(* Logix 5000 project; controller FV vendor 1 type 14 code 217 rev 31.11; software revision 31.00; part 50 of 63 *)
(* tags used below, declared in another part *)
   CheckTimeMask : INT;
   Delphi_Does_Eng_Func : BOOL;
   FV_ALARM : PlantItem;   // ALARM
   FV_AV1 : PlantItem;   // AV1
   FV_AV1A : PlantItem;   // AV1A
   FV_AV2 : PlantItem;   // AV2
   FV_AV3 : PlantItem;   // AV3
   FV_AV4 : PlantItem;   // AV4
   FV_AV4A : PlantItem;   // AV4A
   FV_FV10C : PlantItem;   // FV10C
   FV_FV10J : PlantItem;   // FV10J
   FV_FV11C : PlantItem;   // FV11C
   FV_FV11J : PlantItem;   // FV11J
   FV_FV12C : PlantItem;   // FV12C
   FV_FV12J : PlantItem;   // FV12J
   FV_FV13C : PlantItem;   // FV13C
   FV_FV13J : PlantItem;   // FV13J
   FV_FV14C : PlantItem;   // FV14C
   FV_FV14J : PlantItem;   // FV14J
   FV_FV15C : PlantItem;   // FV15C
   FV_FV15J : PlantItem;   // FV15J
   FV_FV16C : PlantItem;   // FV16C
   FV_FV16J : PlantItem;   // FV16J
   FV_FV17C : PlantItem;   // FV17C
   FV_FV17J : PlantItem;   // FV17J
   FV_FV18C : PlantItem;   // FV18C
   FV_FV18J : PlantItem;   // FV18J
   FV_FV19C : PlantItem;   // FV19C
   FV_FV19J : PlantItem;   // FV19J
   FV_FV20C : PlantItem;   // FV20C
   FV_FV20J : PlantItem;   // FV20J
   FV_FV21C : PlantItem;   // FV21C
   FV_FV21J : PlantItem;   // FV21J
   FV_FV22C : PlantItem;   // FV22C
   FV_FV22J : PlantItem;   // FV22J
   FV_FV23C : PlantItem;   // FV23C
   FV_FV23J : PlantItem;   // FV23J
   FV_FV24C : PlantItem;   // FV24C
   FV_FV24J : PlantItem;   // FV24J
   FV_FV25C : PlantItem;   // FV25C
   FV_FV25J : PlantItem;   // FV25J
   FV_FV26C : PlantItem;   // FV26C
   FV_FV26J : PlantItem;   // FV26J
   FV_FV27C : PlantItem;   // FV27C
   FV_FV27J : PlantItem;   // FV27J
   FV_FV28C : PlantItem;   // FV28C
   FV_FV28J : PlantItem;   // FV28J
   FV_FV29C : PlantItem;   // FV29C
   FV_FV29J : PlantItem;   // FV29J
   FV_FV30C : PlantItem;   // FV30C
   FV_FV30J : PlantItem;   // FV30J
   FV_FV31C : PlantItem;   // FV31C
   FV_FV31J : PlantItem;   // FV31J
   FV_N255 : INT[255];   // Old Checkwords to keep Delphi working in the interim before full changeover.
   FV_PUMP1 : PlantItem;   // PUMP1
   FV_PUMP2 : PlantItem;   // PUMP2
   FV_PUMP3 : PlantItem;   // PUMP3
   FV_R2V1 : PlantItem;   // R2V1
   FV_R2V2 : PlantItem;   // R2V2
   FV_SOV1 : PlantItem;   // SOV1
   FV_SOV2 : PlantItem;   // SOV2
   FV_WYT1R : PlantItem;   // WYT1R
   FV_WYT2R : PlantItem;   // WYT2R
   FV_WYTR1 : PlantItem;   // WYTR1
   FV_WYTR2 : PlantItem;   // WYTR2
   FV_YSV1CV : PlantItem;   // YSV1CV
   FV_YSV1J : PlantItem;   // YSV1J
   FV_YSV1R : PlantItem;   // YSV1R
   FV_YSV2CV : PlantItem;   // YSV2CV
   FV_YSV2J : PlantItem;   // YSV2J
   FV_YSV2O : PlantItem;   // YSV2O
   FV_YSV2R : PlantItem;   // YSV2R
   FV_YSV3J : PlantItem;   // YSV3J
   FV_YSV3O : PlantItem;   // YSV3O
   FV_YSV3R : PlantItem;   // YSV3R
   TempChecktime : DINT;
(* FV_Common, continued *)

   108: XIC(Delphi_Does_Eng_Func)AND(FV_N255[19],CheckTimeMask,TempChecktime)[GRT(TempChecktime,0) DIV(TempChecktime,8,FV_FV10C.CheckTime) ,EQU(TempChecktime,0) OTL(FV_N255[19].6) ];
   109: XIC(Delphi_Does_Eng_Func)AND(FV_N255[20],CheckTimeMask,TempChecktime)[GRT(TempChecktime,0) DIV(TempChecktime,8,FV_FV10J.CheckTime) ,EQU(TempChecktime,0) OTL(FV_N255[20].6) ];
   110: XIC(Delphi_Does_Eng_Func)AND(FV_N255[21],CheckTimeMask,TempChecktime)[GRT(TempChecktime,0) DIV(TempChecktime,8,FV_FV11C.CheckTime) ,EQU(TempChecktime,0) OTL(FV_N255[21].6) ];
   111: XIC(Delphi_Does_Eng_Func)AND(FV_N255[22],CheckTimeMask,TempChecktime)[GRT(TempChecktime,0) DIV(TempChecktime,8,FV_FV11J.CheckTime) ,EQU(TempChecktime,0) OTL(FV_N255[22].6) ];
   112: XIC(Delphi_Does_Eng_Func)AND(FV_N255[23],CheckTimeMask,TempChecktime)[GRT(TempChecktime,0) DIV(TempChecktime,8,FV_FV12C.CheckTime) ,EQU(TempChecktime,0) OTL(FV_N255[23].6) ];
   113: XIC(Delphi_Does_Eng_Func)AND(FV_N255[24],CheckTimeMask,TempChecktime)[GRT(TempChecktime,0) DIV(TempChecktime,8,FV_FV12J.CheckTime) ,EQU(TempChecktime,0) OTL(FV_N255[24].6) ];
   114: XIC(Delphi_Does_Eng_Func)AND(FV_N255[25],CheckTimeMask,TempChecktime)[GRT(TempChecktime,0) DIV(TempChecktime,8,FV_FV13C.CheckTime) ,EQU(TempChecktime,0) OTL(FV_N255[25].6) ];
   115: XIC(Delphi_Does_Eng_Func)AND(FV_N255[26],CheckTimeMask,TempChecktime)[GRT(TempChecktime,0) DIV(TempChecktime,8,FV_FV13J.CheckTime) ,EQU(TempChecktime,0) OTL(FV_N255[26].6) ];
   116: XIC(Delphi_Does_Eng_Func)AND(FV_N255[27],CheckTimeMask,TempChecktime)[GRT(TempChecktime,0) DIV(TempChecktime,8,FV_FV14C.CheckTime) ,EQU(TempChecktime,0) OTL(FV_N255[27].6) ];
   117: XIC(Delphi_Does_Eng_Func)AND(FV_N255[28],CheckTimeMask,TempChecktime)[GRT(TempChecktime,0) DIV(TempChecktime,8,FV_FV14J.CheckTime) ,EQU(TempChecktime,0) OTL(FV_N255[28].6) ];
   118: XIC(Delphi_Does_Eng_Func)AND(FV_N255[29],CheckTimeMask,TempChecktime)[GRT(TempChecktime,0) DIV(TempChecktime,8,FV_FV15C.CheckTime) ,EQU(TempChecktime,0) OTL(FV_N255[29].6) ];
   119: XIC(Delphi_Does_Eng_Func)AND(FV_N255[30],CheckTimeMask,TempChecktime)[GRT(TempChecktime,0) DIV(TempChecktime,8,FV_FV15J.CheckTime) ,EQU(TempChecktime,0) OTL(FV_N255[30].6) ];
   120: XIC(Delphi_Does_Eng_Func)AND(FV_N255[31],CheckTimeMask,TempChecktime)[GRT(TempChecktime,0) DIV(TempChecktime,8,FV_FV16C.CheckTime) ,EQU(TempChecktime,0) OTL(FV_N255[31].6) ];
   121: XIC(Delphi_Does_Eng_Func)AND(FV_N255[32],CheckTimeMask,TempChecktime)[GRT(TempChecktime,0) DIV(TempChecktime,8,FV_FV16J.CheckTime) ,EQU(TempChecktime,0) OTL(FV_N255[32].6) ];
   122: XIC(Delphi_Does_Eng_Func)AND(FV_N255[33],CheckTimeMask,TempChecktime)[GRT(TempChecktime,0) DIV(TempChecktime,8,FV_FV17C.CheckTime) ,EQU(TempChecktime,0) OTL(FV_N255[33].6) ];
   123: XIC(Delphi_Does_Eng_Func)AND(FV_N255[34],CheckTimeMask,TempChecktime)[GRT(TempChecktime,0) DIV(TempChecktime,8,FV_FV17J.CheckTime) ,EQU(TempChecktime,0) OTL(FV_N255[34].6) ];
   124: XIC(Delphi_Does_Eng_Func)AND(FV_N255[35],CheckTimeMask,TempChecktime)[GRT(TempChecktime,0) DIV(TempChecktime,8,FV_FV18C.CheckTime) ,EQU(TempChecktime,0) OTL(FV_N255[35].6) ];
   125: XIC(Delphi_Does_Eng_Func)AND(FV_N255[36],CheckTimeMask,TempChecktime)[GRT(TempChecktime,0) DIV(TempChecktime,8,FV_FV18J.CheckTime) ,EQU(TempChecktime,0) OTL(FV_N255[36].6) ];
   126: XIC(Delphi_Does_Eng_Func)AND(FV_N255[37],CheckTimeMask,TempChecktime)[GRT(TempChecktime,0) DIV(TempChecktime,8,FV_FV19C.CheckTime) ,EQU(TempChecktime,0) OTL(FV_N255[37].6) ];
   127: XIC(Delphi_Does_Eng_Func)AND(FV_N255[38],CheckTimeMask,TempChecktime)[GRT(TempChecktime,0) DIV(TempChecktime,8,FV_FV19J.CheckTime) ,EQU(TempChecktime,0) OTL(FV_N255[38].6) ];
   128: XIC(Delphi_Does_Eng_Func)AND(FV_N255[39],CheckTimeMask,TempChecktime)[GRT(TempChecktime,0) DIV(TempChecktime,8,FV_FV20C.CheckTime) ,EQU(TempChecktime,0) OTL(FV_N255[39].6) ];
   129: XIC(Delphi_Does_Eng_Func)AND(FV_N255[40],CheckTimeMask,TempChecktime)[GRT(TempChecktime,0) DIV(TempChecktime,8,FV_FV20J.CheckTime) ,EQU(TempChecktime,0) OTL(FV_N255[40].6) ];
   130: XIC(Delphi_Does_Eng_Func)AND(FV_N255[41],CheckTimeMask,TempChecktime)[GRT(TempChecktime,0) DIV(TempChecktime,8,FV_FV21C.CheckTime) ,EQU(TempChecktime,0) OTL(FV_N255[41].6) ];
   131: XIC(Delphi_Does_Eng_Func)AND(FV_N255[42],CheckTimeMask,TempChecktime)[GRT(TempChecktime,0) DIV(TempChecktime,8,FV_FV21J.CheckTime) ,EQU(TempChecktime,0) OTL(FV_N255[42].6) ];
   132: XIC(Delphi_Does_Eng_Func)AND(FV_N255[43],CheckTimeMask,TempChecktime)[GRT(TempChecktime,0) DIV(TempChecktime,8,FV_FV22C.CheckTime) ,EQU(TempChecktime,0) OTL(FV_N255[43].6) ];
   133: XIC(Delphi_Does_Eng_Func)AND(FV_N255[44],CheckTimeMask,TempChecktime)[GRT(TempChecktime,0) DIV(TempChecktime,8,FV_FV22J.CheckTime) ,EQU(TempChecktime,0) OTL(FV_N255[44].6) ];
   134: XIC(Delphi_Does_Eng_Func)AND(FV_N255[45],CheckTimeMask,TempChecktime)[GRT(TempChecktime,0) DIV(TempChecktime,8,FV_FV23C.CheckTime) ,EQU(TempChecktime,0) OTL(FV_N255[45].6) ];
   135: XIC(Delphi_Does_Eng_Func)AND(FV_N255[46],CheckTimeMask,TempChecktime)[GRT(TempChecktime,0) DIV(TempChecktime,8,FV_FV23J.CheckTime) ,EQU(TempChecktime,0) OTL(FV_N255[46].6) ];
   136: XIC(Delphi_Does_Eng_Func)AND(FV_N255[47],CheckTimeMask,TempChecktime)[GRT(TempChecktime,0) DIV(TempChecktime,8,FV_FV24C.CheckTime) ,EQU(TempChecktime,0) OTL(FV_N255[47].6) ];
   137: XIC(Delphi_Does_Eng_Func)AND(FV_N255[48],CheckTimeMask,TempChecktime)[GRT(TempChecktime,0) DIV(TempChecktime,8,FV_FV24J.CheckTime) ,EQU(TempChecktime,0) OTL(FV_N255[48].6) ];
   138: XIC(Delphi_Does_Eng_Func)AND(FV_N255[49],CheckTimeMask,TempChecktime)[GRT(TempChecktime,0) DIV(TempChecktime,8,FV_FV25C.CheckTime) ,EQU(TempChecktime,0) OTL(FV_N255[49].6) ];
   139: XIC(Delphi_Does_Eng_Func)AND(FV_N255[50],CheckTimeMask,TempChecktime)[GRT(TempChecktime,0) DIV(TempChecktime,8,FV_FV25J.CheckTime) ,EQU(TempChecktime,0) OTL(FV_N255[50].6) ];
   140: XIC(Delphi_Does_Eng_Func)AND(FV_N255[53],CheckTimeMask,TempChecktime)[GRT(TempChecktime,0) DIV(TempChecktime,8,FV_YSV2O.CheckTime) ,EQU(TempChecktime,0) OTL(FV_N255[53].6) ];
   141: XIC(Delphi_Does_Eng_Func)AND(FV_N255[54],CheckTimeMask,TempChecktime)[GRT(TempChecktime,0) DIV(TempChecktime,8,FV_ALARM.CheckTime) ,EQU(TempChecktime,0) OTL(FV_N255[54].6) ];
   142: XIC(Delphi_Does_Eng_Func)AND(FV_N255[55],CheckTimeMask,TempChecktime)[GRT(TempChecktime,0) DIV(TempChecktime,8,FV_YSV3O.CheckTime) ,EQU(TempChecktime,0) OTL(FV_N255[55].6) ];
   143: XIC(Delphi_Does_Eng_Func)AND(FV_N255[56],CheckTimeMask,TempChecktime)[GRT(TempChecktime,0) DIV(TempChecktime,8,FV_YSV3J.CheckTime) ,EQU(TempChecktime,0) OTL(FV_N255[56].6) ];
   144: XIC(Delphi_Does_Eng_Func)AND(FV_N255[57],CheckTimeMask,TempChecktime)[GRT(TempChecktime,0) DIV(TempChecktime,8,FV_YSV3R.CheckTime) ,EQU(TempChecktime,0) OTL(FV_N255[57].6) ];
   145: XIC(Delphi_Does_Eng_Func)AND(FV_N255[58],CheckTimeMask,TempChecktime)[GRT(TempChecktime,0) DIV(TempChecktime,8,FV_YSV1J.CheckTime) ,EQU(TempChecktime,0) OTL(FV_N255[58].6) ];
   146: XIC(Delphi_Does_Eng_Func)AND(FV_N255[60],CheckTimeMask,TempChecktime)[GRT(TempChecktime,0) DIV(TempChecktime,8,FV_YSV2J.CheckTime) ,EQU(TempChecktime,0) OTL(FV_N255[60].6) ];
   147: XIC(Delphi_Does_Eng_Func)AND(FV_N255[61],CheckTimeMask,TempChecktime)[GRT(TempChecktime,0) DIV(TempChecktime,8,FV_YSV2R.CheckTime) ,EQU(TempChecktime,0) OTL(FV_N255[61].6) ];
   148: XIC(Delphi_Does_Eng_Func)AND(FV_N255[62],CheckTimeMask,TempChecktime)[GRT(TempChecktime,0) DIV(TempChecktime,8,FV_PUMP1.CheckTime) ,EQU(TempChecktime,0) OTL(FV_N255[62].6) ];
   149: XIC(Delphi_Does_Eng_Func)AND(FV_N255[63],CheckTimeMask,TempChecktime)[GRT(TempChecktime,0) DIV(TempChecktime,8,FV_PUMP2.CheckTime) ,EQU(TempChecktime,0) OTL(FV_N255[63].6) ];
   150: XIC(Delphi_Does_Eng_Func)AND(FV_N255[64],CheckTimeMask,TempChecktime)[GRT(TempChecktime,0) DIV(TempChecktime,8,FV_PUMP3.CheckTime) ,EQU(TempChecktime,0) OTL(FV_N255[64].6) ];
   151: XIC(Delphi_Does_Eng_Func)AND(FV_N255[71],CheckTimeMask,TempChecktime)[GRT(TempChecktime,0) DIV(TempChecktime,8,FV_SOV1.CheckTime) ,EQU(TempChecktime,0) OTL(FV_N255[71].6) ];
   152: XIC(Delphi_Does_Eng_Func)AND(FV_N255[72],CheckTimeMask,TempChecktime)[GRT(TempChecktime,0) DIV(TempChecktime,8,FV_SOV2.CheckTime) ,EQU(TempChecktime,0) OTL(FV_N255[72].6) ];
   153: XIC(Delphi_Does_Eng_Func)AND(FV_N255[77],CheckTimeMask,TempChecktime)[GRT(TempChecktime,0) DIV(TempChecktime,8,FV_YSV1CV.CheckTime) ,EQU(TempChecktime,0) OTL(FV_N255[77].6) ];
   154: XIC(Delphi_Does_Eng_Func)AND(FV_N255[78],CheckTimeMask,TempChecktime)[GRT(TempChecktime,0) DIV(TempChecktime,8,FV_YSV2CV.CheckTime) ,EQU(TempChecktime,0) OTL(FV_N255[78].6) ];
   155: XIC(Delphi_Does_Eng_Func)AND(FV_N255[81],CheckTimeMask,TempChecktime)[GRT(TempChecktime,0) DIV(TempChecktime,8,FV_FV26J.CheckTime) ,EQU(TempChecktime,0) OTL(FV_N255[81].6) ];
   156: XIC(Delphi_Does_Eng_Func)AND(FV_N255[82],CheckTimeMask,TempChecktime)[GRT(TempChecktime,0) DIV(TempChecktime,8,FV_FV26C.CheckTime) ,EQU(TempChecktime,0) OTL(FV_N255[82].6) ];
   157: XIC(Delphi_Does_Eng_Func)AND(FV_N255[83],CheckTimeMask,TempChecktime)[GRT(TempChecktime,0) DIV(TempChecktime,8,FV_FV27J.CheckTime) ,EQU(TempChecktime,0) OTL(FV_N255[83].6) ];
   158: XIC(Delphi_Does_Eng_Func)AND(FV_N255[84],CheckTimeMask,TempChecktime)[GRT(TempChecktime,0) DIV(TempChecktime,8,FV_FV27C.CheckTime) ,EQU(TempChecktime,0) OTL(FV_N255[84].6) ];
   159: XIC(Delphi_Does_Eng_Func)AND(FV_N255[85],CheckTimeMask,TempChecktime)[GRT(TempChecktime,0) DIV(TempChecktime,8,FV_FV28J.CheckTime) ,EQU(TempChecktime,0) OTL(FV_N255[85].6) ];
   160: XIC(Delphi_Does_Eng_Func)AND(FV_N255[86],CheckTimeMask,TempChecktime)[GRT(TempChecktime,0) DIV(TempChecktime,8,FV_FV28C.CheckTime) ,EQU(TempChecktime,0) OTL(FV_N255[86].6) ];
   161: XIC(Delphi_Does_Eng_Func)AND(FV_N255[87],CheckTimeMask,TempChecktime)[GRT(TempChecktime,0) DIV(TempChecktime,8,FV_FV29J.CheckTime) ,EQU(TempChecktime,0) OTL(FV_N255[87].6) ];
   162: XIC(Delphi_Does_Eng_Func)AND(FV_N255[88],CheckTimeMask,TempChecktime)[GRT(TempChecktime,0) DIV(TempChecktime,8,FV_FV29C.CheckTime) ,EQU(TempChecktime,0) OTL(FV_N255[88].6) ];
   163: XIC(Delphi_Does_Eng_Func)AND(FV_N255[89],CheckTimeMask,TempChecktime)[GRT(TempChecktime,0) DIV(TempChecktime,8,FV_FV30J.CheckTime) ,EQU(TempChecktime,0) OTL(FV_N255[89].6) ];
   164: XIC(Delphi_Does_Eng_Func)AND(FV_N255[90],CheckTimeMask,TempChecktime)[GRT(TempChecktime,0) DIV(TempChecktime,8,FV_FV30C.CheckTime) ,EQU(TempChecktime,0) OTL(FV_N255[90].6) ];
   165: XIC(Delphi_Does_Eng_Func)AND(FV_N255[91],CheckTimeMask,TempChecktime)[GRT(TempChecktime,0) DIV(TempChecktime,8,FV_FV31J.CheckTime) ,EQU(TempChecktime,0) OTL(FV_N255[91].6) ];
   166: XIC(Delphi_Does_Eng_Func)AND(FV_N255[92],CheckTimeMask,TempChecktime)[GRT(TempChecktime,0) DIV(TempChecktime,8,FV_FV31C.CheckTime) ,EQU(TempChecktime,0) OTL(FV_N255[92].6) ];
   167: XIC(Delphi_Does_Eng_Func)AND(FV_N255[79],CheckTimeMask,TempChecktime)[GRT(TempChecktime,0) DIV(TempChecktime,8,FV_WYT1R.CheckTime) ,EQU(TempChecktime,0) OTL(FV_N255[79].6) ];
   168: XIC(Delphi_Does_Eng_Func)AND(FV_N255[80],CheckTimeMask,TempChecktime)[GRT(TempChecktime,0) DIV(TempChecktime,8,FV_WYT2R.CheckTime) ,EQU(TempChecktime,0) OTL(FV_N255[80].6) ];
   169: XIC(Delphi_Does_Eng_Func)AND(FV_N255[59],CheckTimeMask,TempChecktime)[GRT(TempChecktime,0) DIV(TempChecktime,8,FV_YSV1R.CheckTime) ,EQU(TempChecktime,0) OTL(FV_N255[59].6) ];
   170: XIC(Delphi_Does_Eng_Func)AND(FV_N255[65],CheckTimeMask,TempChecktime)[GRT(TempChecktime,0) DIV(TempChecktime,8,FV_AV1.CheckTime) ,EQU(TempChecktime,0) OTL(FV_N255[65].6) ];
   171: XIC(Delphi_Does_Eng_Func)AND(FV_N255[66],CheckTimeMask,TempChecktime)[GRT(TempChecktime,0) DIV(TempChecktime,8,FV_AV2.CheckTime) ,EQU(TempChecktime,0) OTL(FV_N255[66].6) ];
   172: XIC(Delphi_Does_Eng_Func)AND(FV_N255[67],CheckTimeMask,TempChecktime)[GRT(TempChecktime,0) DIV(TempChecktime,8,FV_AV3.CheckTime) ,EQU(TempChecktime,0) OTL(FV_N255[67].6) ];
   173: XIC(Delphi_Does_Eng_Func)AND(FV_N255[68],CheckTimeMask,TempChecktime)[GRT(TempChecktime,0) DIV(TempChecktime,8,FV_AV4.CheckTime) ,EQU(TempChecktime,0) OTL(FV_N255[68].6) ];
   174: XIC(Delphi_Does_Eng_Func)AND(FV_N255[69],CheckTimeMask,TempChecktime)[GRT(TempChecktime,0) DIV(TempChecktime,8,FV_AV1A.CheckTime) ,EQU(TempChecktime,0) OTL(FV_N255[69].6) ];
   175: XIC(Delphi_Does_Eng_Func)AND(FV_N255[70],CheckTimeMask,TempChecktime)[GRT(TempChecktime,0) DIV(TempChecktime,8,FV_AV4A.CheckTime) ,EQU(TempChecktime,0) OTL(FV_N255[70].6) ];
   176: XIC(Delphi_Does_Eng_Func)AND(FV_N255[73],CheckTimeMask,TempChecktime)[GRT(TempChecktime,0) DIV(TempChecktime,8,FV_WYTR1.CheckTime) ,EQU(TempChecktime,0) OTL(FV_N255[73].6) ];
   177: XIC(Delphi_Does_Eng_Func)AND(FV_N255[74],CheckTimeMask,TempChecktime)[GRT(TempChecktime,0) DIV(TempChecktime,8,FV_WYTR2.CheckTime) ,EQU(TempChecktime,0) OTL(FV_N255[74].6) ];
   178: XIC(Delphi_Does_Eng_Func)AND(FV_N255[75],CheckTimeMask,TempChecktime)[GRT(TempChecktime,0) DIV(TempChecktime,8,FV_R2V1.CheckTime) ,EQU(TempChecktime,0) OTL(FV_N255[75].6) ];
   179: XIC(Delphi_Does_Eng_Func)AND(FV_N255[76],CheckTimeMask,TempChecktime)[GRT(TempChecktime,0) DIV(TempChecktime,8,FV_R2V2.CheckTime) ,EQU(TempChecktime,0) OTL(FV_N255[76].6) ];
END_ROUTINE
